REGION Network 28 (STL): spare- VB chan 8
         A     "Epics_to_PLC"."spare-VB-8".cmdSet;
         S     "voie 8 chaufferette BV";
         A     "Epics_to_PLC"."spare-VB-8".cmdRst;
         R     "voie 8 chaufferette BV";
END_REGION

REGION Network 29 (STL): spare- VB chan 9
         A     "Epics_to_PLC"."spare-VB-9".cmdSet;
         S     "voie 9 chaufferette BV";
         A     "Epics_to_PLC"."spare-VB-9".cmdRst;
         R     "voie 9 chaufferette BV";
END_REGION

REGION Network 30 (STL): spare- VB chan 10
         A     "Epics_to_PLC"."spare-VB-10".cmdSet;
         S     "voie 10  chaufferette BV";
         A     "Epics_to_PLC"."spare-VB-10".cmdRst;
         R     "voie 10  chaufferette BV";
END_REGION

REGION Network 31 (STL): spare - VB chan 11
         A     "Epics_to_PLC"."spare-VB-11".cmdSet;
         S     "voie 11 chaufferette BV";
         A     "Epics_to_PLC"."spare-VB-11".cmdRst;
         R     "voie 11 chaufferette BV";
END_REGION

REGION Network 32 (STL): spare - CM chan 5
         A     "Epics_to_PLC"."spare-CM-5".cmdSet;
         S     "voie 5 chaufferette CM";
         A     "Epics_to_PLC"."spare-CM-5".cmdRst;
         R     "voie 5 chaufferette CM";
END_REGION

REGION Network 33 (STL): spare - CM chan 6
         A     "Epics_to_PLC"."spare-CM-6".cmdSet;
         S     "voie 6 chaufferette CM";
         A     "Epics_to_PLC"."spare-CM-6".cmdRst;
         R     "voie 6 chaufferette CM";
END_REGION

REGION Network 34 (STL): spare - CM chan 7
         A     "Epics_to_PLC"."spare-CM-7".cmdSet;
         S     "voie 7 chaufferette CM";
         A     "Epics_to_PLC"."spare-CM-7".cmdRst;
         R     "voie 7 chaufferette CM";
END_REGION

REGION Network 35 (STL): spare - CM chan 8
         A     "Epics_to_PLC"."spare-CM-8".cmdSet;
         S     "voie 8 chaufferette CM";
         A     "Epics_to_PLC"."spare-CM-8".cmdRst;
         R     "voie 8 chaufferette CM";
END_REGION

REGION Network 36 (STL): spare - CM chan 10
         A     "Epics_to_PLC"."spare-CM-10".cmdSet;
         S     "voie 10 chaufferette CM";
         A     "Epics_to_PLC"."spare-CM-10".cmdRst;
         R     "voie 10 chaufferette CM";
END_REGION

REGION Network 37 (STL): spare - CM chan 12
         A     "Epics_to_PLC"."spare-CM-12".cmdSet;
         S     "voie 12 chaufferette CM";
         A     "Epics_to_PLC"."spare-CM-12".cmdRst;
         R     "voie 12 chaufferette CM";
END_REGION

REGION Network 38 (STL): Bit commands
         A     "Epics_to_PLC".cmdAutoMode;
         R     "Graph/manuelle";
         A     "Epics_to_PLC".cmdManMode;
         S     "Graph/manuelle";
         A     "Epics_to_PLC".cmdGrafcetInit;
         =     "MettreEtatInitial";
         A     "Epics_to_PLC".cmdGrafcetErrRst;
         =     "AcquitterErreurGraph";
         A     "Epics_to_PLC".cmdStartConditioning;
         =     "CmdVanneEtatCdt";
         A     "Epics_to_PLC".cmdCondOK;
         =     "CdtInfraOk";
         A     "Epics_to_PLC".cmdCondERR;
         =     "CdtInfraErreur";
         A     "Epics_to_PLC".cmdStartLN2cooling;
         =     "DmdMefAzote";
         A     "Epics_to_PLC".cmdStartLHecooling;
         =     "DmdMefHelium";
         A     "Epics_to_PLC".cmdStart2Kmode;
         =     "DmdMode2K";
         A     "Epics_to_PLC".cmdStop2Kmode;
         =     "DmdArretMode2k";
         A     "Epics_to_PLC".cmdStartSTBYmode;
         =     "DmdModeStandby";
         A     "Epics_to_PLC".cmdStopSTBYmode;
         =     "DmdArretModeStandby";
         A     "Epics_to_PLC".cmdStartHeating;
         =     "StartHeating";
         A     "Epics_to_PLC".cmdStopHeating;
         =     "StopHeating";
         A     "Epics_to_PLC".cmdSelLT01;
         R     "LT_CM".LT02_selCtrl;
         A     "Epics_to_PLC".cmdSelLT02;
         S     "LT_CM".LT02_selCtrl;
END_REGION

REGION Network 39: Real parameters (LHe level PIDs settings)
   RUNG wire#powerrail
      Contact( "Epics_to_PLC".TrigPID_CV01.cmdSet )
      { S7_GenerateENO := "TRUE" } Move(in := "Epics_to_PLC".TrigPID_CV01.cSetV, out1 => "TriggerPIDcv01")
      { S7_GenerateENO := "TRUE" } Move(in := "Epics_to_PLC".TrigPID_CV01.cSetV, out1 => "S8_parameters".TrigPID_CV01)
      R_Coil( "Epics_to_PLC".TrigPID_CV01.cmdSet )
   END_RUNG
   // the same network as SCL:
   // ENO of a box is taken as its EN; it also drops when the box reports an error
   IF "Epics_to_PLC".TrigPID_CV01.cmdSet THEN
       "TriggerPIDcv01" := "Epics_to_PLC".TrigPID_CV01.cSetV;
       "S8_parameters".TrigPID_CV01 := "Epics_to_PLC".TrigPID_CV01.cSetV;
       "Epics_to_PLC".TrigPID_CV01.cmdSet := FALSE;
   END_IF;
END_REGION

REGION Network 40: Real parameters (LHe level PIDs settings)
   RUNG wire#powerrail
      Contact( "Epics_to_PLC".TrigPID_CV02.cmdSet )
      { S7_GenerateENO := "TRUE" } Move(in := "Epics_to_PLC".TrigPID_CV02.cSetV, out1 => "TriggerPIDcv02")
      { S7_GenerateENO := "TRUE" } Move(in := "Epics_to_PLC".TrigPID_CV02.cSetV, out1 => "S6_parameters".TrigPID_CV02)
      R_Coil( "Epics_to_PLC".TrigPID_CV02.cmdSet )
   END_RUNG
   // the same network as SCL:
   // ENO of a box is taken as its EN; it also drops when the box reports an error
   IF "Epics_to_PLC".TrigPID_CV02.cmdSet THEN
       "TriggerPIDcv02" := "Epics_to_PLC".TrigPID_CV02.cSetV;
       "S6_parameters".TrigPID_CV02 := "Epics_to_PLC".TrigPID_CV02.cSetV;
       "Epics_to_PLC".TrigPID_CV02.cmdSet := FALSE;
   END_IF;
END_REGION

REGION Network 41: Real parameters (LHe level PIDs settings)
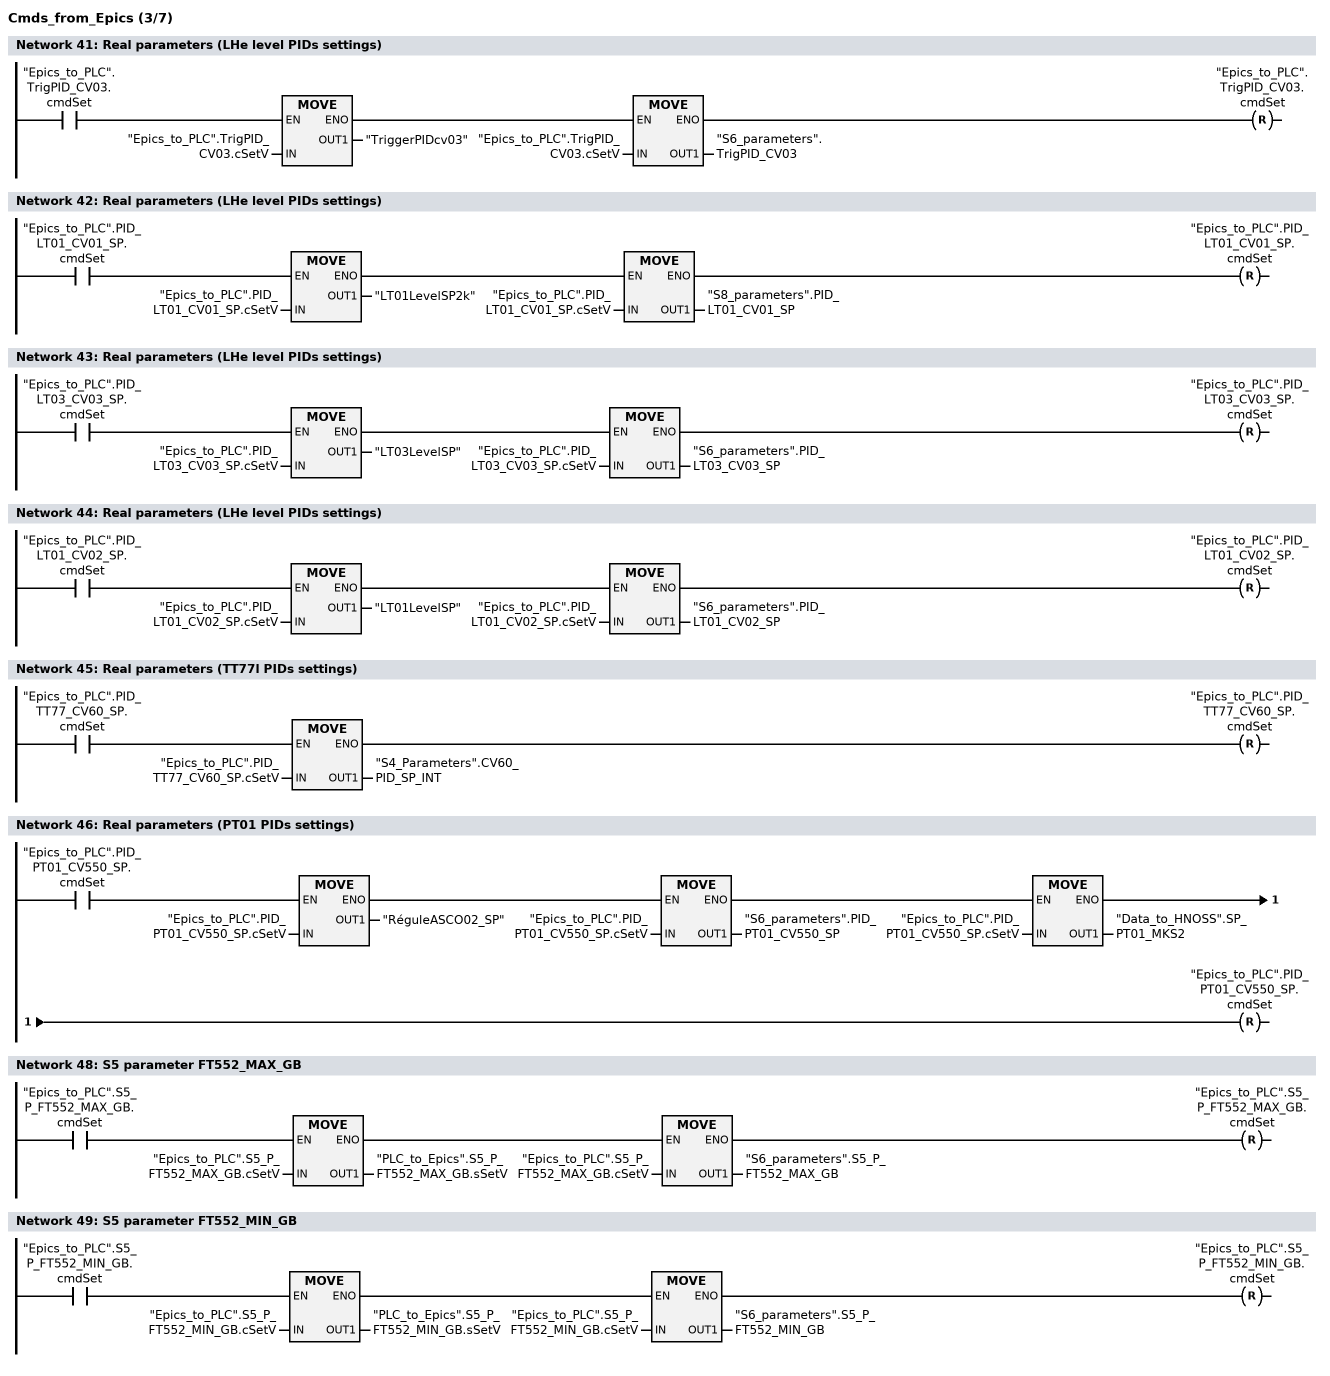
   RUNG wire#powerrail
      Contact( "Epics_to_PLC".TrigPID_CV03.cmdSet )
      { S7_GenerateENO := "TRUE" } Move(in := "Epics_to_PLC".TrigPID_CV03.cSetV, out1 => "TriggerPIDcv03")
      { S7_GenerateENO := "TRUE" } Move(in := "Epics_to_PLC".TrigPID_CV03.cSetV, out1 => "S6_parameters".TrigPID_CV03)
      R_Coil( "Epics_to_PLC".TrigPID_CV03.cmdSet )
   END_RUNG
   // the same network as SCL:
   // ENO of a box is taken as its EN; it also drops when the box reports an error
   IF "Epics_to_PLC".TrigPID_CV03.cmdSet THEN
       "TriggerPIDcv03" := "Epics_to_PLC".TrigPID_CV03.cSetV;
       "S6_parameters".TrigPID_CV03 := "Epics_to_PLC".TrigPID_CV03.cSetV;
       "Epics_to_PLC".TrigPID_CV03.cmdSet := FALSE;
   END_IF;
END_REGION

REGION Network 42: Real parameters (LHe level PIDs settings)
   RUNG wire#powerrail
      Contact( "Epics_to_PLC".PID_LT01_CV01_SP.cmdSet )
      { S7_GenerateENO := "TRUE" } Move(in := "Epics_to_PLC".PID_LT01_CV01_SP.cSetV, out1 => "LT01LevelSP2k")
      { S7_GenerateENO := "TRUE" } Move(in := "Epics_to_PLC".PID_LT01_CV01_SP.cSetV, out1 => "S8_parameters".PID_LT01_CV01_SP)
      R_Coil( "Epics_to_PLC".PID_LT01_CV01_SP.cmdSet )
   END_RUNG
   // the same network as SCL:
   // ENO of a box is taken as its EN; it also drops when the box reports an error
   IF "Epics_to_PLC".PID_LT01_CV01_SP.cmdSet THEN
       "LT01LevelSP2k" := "Epics_to_PLC".PID_LT01_CV01_SP.cSetV;
       "S8_parameters".PID_LT01_CV01_SP := "Epics_to_PLC".PID_LT01_CV01_SP.cSetV;
       "Epics_to_PLC".PID_LT01_CV01_SP.cmdSet := FALSE;
   END_IF;
END_REGION

REGION Network 43: Real parameters (LHe level PIDs settings)
   RUNG wire#powerrail
      Contact( "Epics_to_PLC".PID_LT03_CV03_SP.cmdSet )
      { S7_GenerateENO := "TRUE" } Move(in := "Epics_to_PLC".PID_LT03_CV03_SP.cSetV, out1 => "LT03LevelSP")
      { S7_GenerateENO := "TRUE" } Move(in := "Epics_to_PLC".PID_LT03_CV03_SP.cSetV, out1 => "S6_parameters".PID_LT03_CV03_SP)
      R_Coil( "Epics_to_PLC".PID_LT03_CV03_SP.cmdSet )
   END_RUNG
   // the same network as SCL:
   // ENO of a box is taken as its EN; it also drops when the box reports an error
   IF "Epics_to_PLC".PID_LT03_CV03_SP.cmdSet THEN
       "LT03LevelSP" := "Epics_to_PLC".PID_LT03_CV03_SP.cSetV;
       "S6_parameters".PID_LT03_CV03_SP := "Epics_to_PLC".PID_LT03_CV03_SP.cSetV;
       "Epics_to_PLC".PID_LT03_CV03_SP.cmdSet := FALSE;
   END_IF;
END_REGION

REGION Network 44: Real parameters (LHe level PIDs settings)
   RUNG wire#powerrail
      Contact( "Epics_to_PLC".PID_LT01_CV02_SP.cmdSet )
      { S7_GenerateENO := "TRUE" } Move(in := "Epics_to_PLC".PID_LT01_CV02_SP.cSetV, out1 => "LT01LevelSP")
      { S7_GenerateENO := "TRUE" } Move(in := "Epics_to_PLC".PID_LT01_CV02_SP.cSetV, out1 => "S6_parameters".PID_LT01_CV02_SP)
      R_Coil( "Epics_to_PLC".PID_LT01_CV02_SP.cmdSet )
   END_RUNG
   // the same network as SCL:
   // ENO of a box is taken as its EN; it also drops when the box reports an error
   IF "Epics_to_PLC".PID_LT01_CV02_SP.cmdSet THEN
       "LT01LevelSP" := "Epics_to_PLC".PID_LT01_CV02_SP.cSetV;
       "S6_parameters".PID_LT01_CV02_SP := "Epics_to_PLC".PID_LT01_CV02_SP.cSetV;
       "Epics_to_PLC".PID_LT01_CV02_SP.cmdSet := FALSE;
   END_IF;
END_REGION

REGION Network 45: Real parameters (TT77l PIDs settings)
   RUNG wire#powerrail
      Contact( "Epics_to_PLC".PID_TT77_CV60_SP.cmdSet )
      { S7_GenerateENO := "TRUE" } Move(in := "Epics_to_PLC".PID_TT77_CV60_SP.cSetV, out1 => "S4_Parameters".CV60_PID_SP_INT)
      R_Coil( "Epics_to_PLC".PID_TT77_CV60_SP.cmdSet )
   END_RUNG
   // the same network as SCL:
   // ENO of a box is taken as its EN; it also drops when the box reports an error
   IF "Epics_to_PLC".PID_TT77_CV60_SP.cmdSet THEN
       "S4_Parameters".CV60_PID_SP_INT := "Epics_to_PLC".PID_TT77_CV60_SP.cSetV;
       "Epics_to_PLC".PID_TT77_CV60_SP.cmdSet := FALSE;
   END_IF;
END_REGION

REGION Network 46: Real parameters (PT01 PIDs settings)
   RUNG wire#powerrail
      Contact( "Epics_to_PLC".PID_PT01_CV550_SP.cmdSet )
      { S7_GenerateENO := "TRUE" } Move(in := "Epics_to_PLC".PID_PT01_CV550_SP.cSetV, out1 => "RéguleASCO02_SP")
      { S7_GenerateENO := "TRUE" } Move(in := "Epics_to_PLC".PID_PT01_CV550_SP.cSetV, out1 => "S6_parameters".PID_PT01_CV550_SP)
      { S7_GenerateENO := "TRUE" } Move(in := "Epics_to_PLC".PID_PT01_CV550_SP.cSetV, out1 => "Data_to_HNOSS".SP_PT01_MKS2)
      R_Coil( "Epics_to_PLC".PID_PT01_CV550_SP.cmdSet )
   END_RUNG
   // the same network as SCL:
   // ENO of a box is taken as its EN; it also drops when the box reports an error
   IF "Epics_to_PLC".PID_PT01_CV550_SP.cmdSet THEN
       "RéguleASCO02_SP" := "Epics_to_PLC".PID_PT01_CV550_SP.cSetV;
       "S6_parameters".PID_PT01_CV550_SP := "Epics_to_PLC".PID_PT01_CV550_SP.cSetV;
       "Data_to_HNOSS".SP_PT01_MKS2 := "Epics_to_PLC".PID_PT01_CV550_SP.cSetV;
       "Epics_to_PLC".PID_PT01_CV550_SP.cmdSet := FALSE;
   END_IF;
END_REGION

REGION Network 47 (STL): Temperatures fromKeithley
         L     "Epics_to_PLC".TTxx;
         T     "ReceivePT100"."TTxx_(K)";
         L     "Epics_to_PLC".TTyy;
         T     "ReceivePT100"."TTyy_(K)";
END_REGION

REGION Network 48: S5 parameter FT552_MAX_GB
   RUNG wire#powerrail
      Contact( "Epics_to_PLC".S5_P_FT552_MAX_GB.cmdSet )
      { S7_GenerateENO := "TRUE" } Move(in := "Epics_to_PLC".S5_P_FT552_MAX_GB.cSetV, out1 => "PLC_to_Epics".S5_P_FT552_MAX_GB.sSetV)
      { S7_GenerateENO := "TRUE" } Move(in := "Epics_to_PLC".S5_P_FT552_MAX_GB.cSetV, out1 => "S6_parameters".S5_P_FT552_MAX_GB)
      R_Coil( "Epics_to_PLC".S5_P_FT552_MAX_GB.cmdSet )
   END_RUNG
   // the same network as SCL:
   // ENO of a box is taken as its EN; it also drops when the box reports an error
   IF "Epics_to_PLC".S5_P_FT552_MAX_GB.cmdSet THEN
       "PLC_to_Epics".S5_P_FT552_MAX_GB.sSetV := "Epics_to_PLC".S5_P_FT552_MAX_GB.cSetV;
       "S6_parameters".S5_P_FT552_MAX_GB := "Epics_to_PLC".S5_P_FT552_MAX_GB.cSetV;
       "Epics_to_PLC".S5_P_FT552_MAX_GB.cmdSet := FALSE;
   END_IF;
END_REGION

REGION Network 49: S5 parameter FT552_MIN_GB
   RUNG wire#powerrail
      Contact( "Epics_to_PLC".S5_P_FT552_MIN_GB.cmdSet )
      { S7_GenerateENO := "TRUE" } Move(in := "Epics_to_PLC".S5_P_FT552_MIN_GB.cSetV, out1 => "PLC_to_Epics".S5_P_FT552_MIN_GB.sSetV)
      { S7_GenerateENO := "TRUE" } Move(in := "Epics_to_PLC".S5_P_FT552_MIN_GB.cSetV, out1 => "S6_parameters".S5_P_FT552_MIN_GB)
      R_Coil( "Epics_to_PLC".S5_P_FT552_MIN_GB.cmdSet )
   END_RUNG
   // the same network as SCL:
   // ENO of a box is taken as its EN; it also drops when the box reports an error
   IF "Epics_to_PLC".S5_P_FT552_MIN_GB.cmdSet THEN
       "PLC_to_Epics".S5_P_FT552_MIN_GB.sSetV := "Epics_to_PLC".S5_P_FT552_MIN_GB.cSetV;
       "S6_parameters".S5_P_FT552_MIN_GB := "Epics_to_PLC".S5_P_FT552_MIN_GB.cSetV;
       "Epics_to_PLC".S5_P_FT552_MIN_GB.cmdSet := FALSE;
   END_IF;
END_REGION

REGION Network 50: S5 parameter FT552_MAX_C
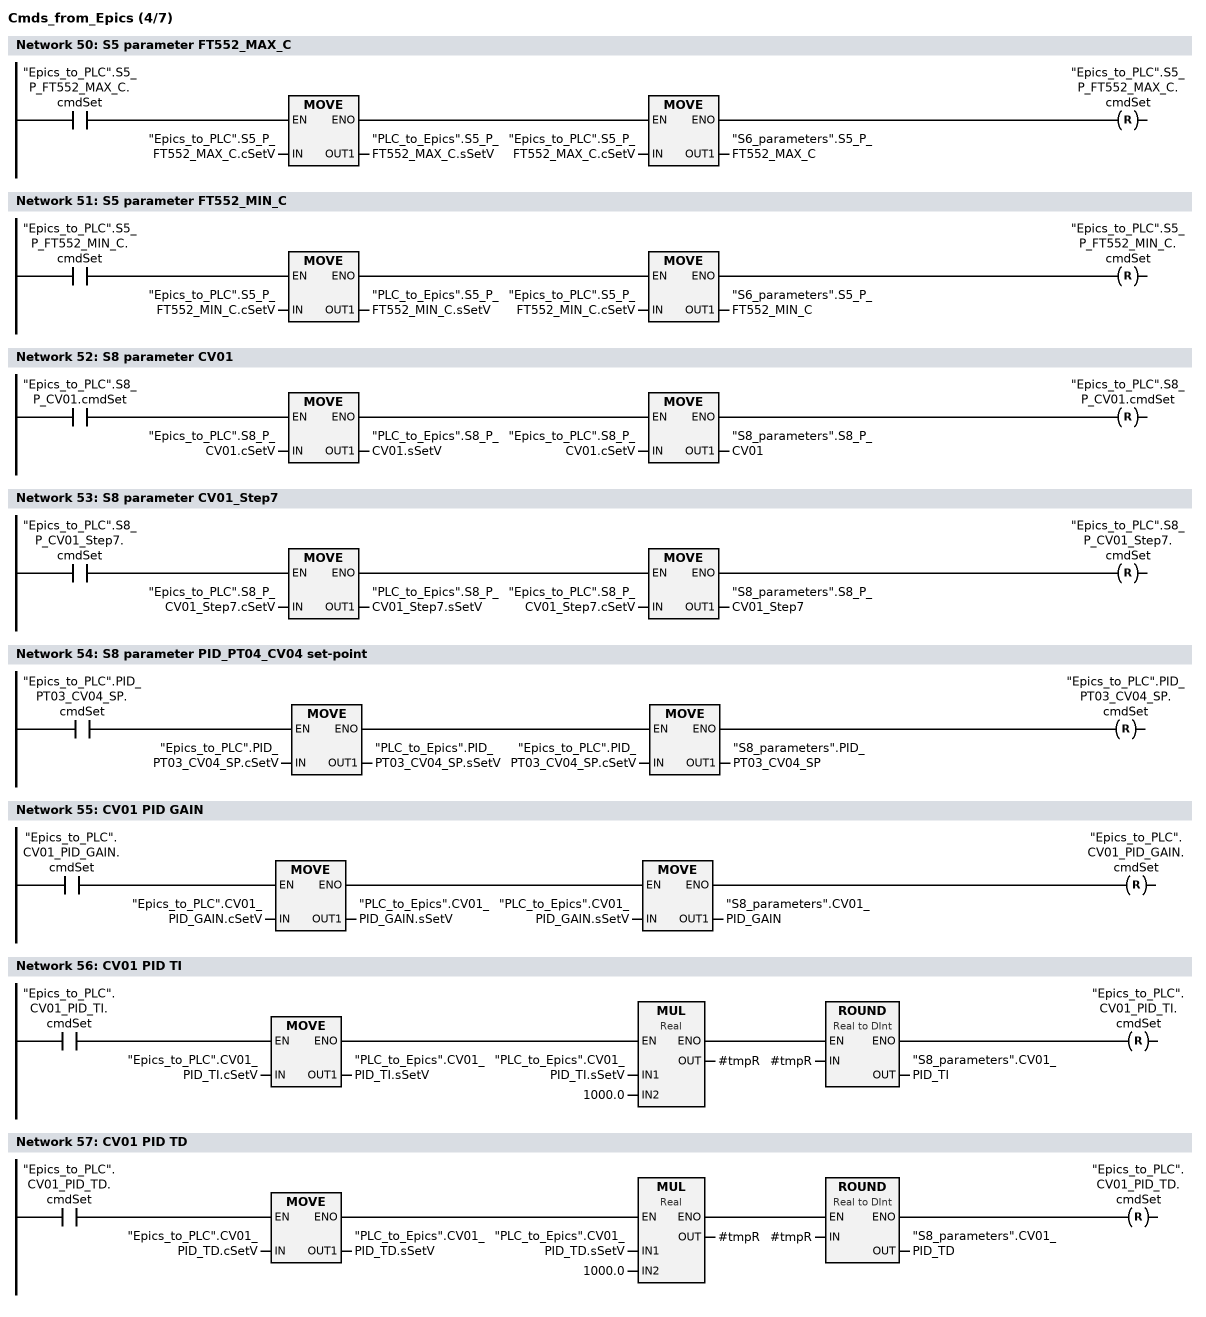
   RUNG wire#powerrail
      Contact( "Epics_to_PLC".S5_P_FT552_MAX_C.cmdSet )
      { S7_GenerateENO := "TRUE" } Move(in := "Epics_to_PLC".S5_P_FT552_MAX_C.cSetV, out1 => "PLC_to_Epics".S5_P_FT552_MAX_C.sSetV)
      { S7_GenerateENO := "TRUE" } Move(in := "Epics_to_PLC".S5_P_FT552_MAX_C.cSetV, out1 => "S6_parameters".S5_P_FT552_MAX_C)
      R_Coil( "Epics_to_PLC".S5_P_FT552_MAX_C.cmdSet )
   END_RUNG
   // the same network as SCL:
   // ENO of a box is taken as its EN; it also drops when the box reports an error
   IF "Epics_to_PLC".S5_P_FT552_MAX_C.cmdSet THEN
       "PLC_to_Epics".S5_P_FT552_MAX_C.sSetV := "Epics_to_PLC".S5_P_FT552_MAX_C.cSetV;
       "S6_parameters".S5_P_FT552_MAX_C := "Epics_to_PLC".S5_P_FT552_MAX_C.cSetV;
       "Epics_to_PLC".S5_P_FT552_MAX_C.cmdSet := FALSE;
   END_IF;
END_REGION

REGION Network 51: S5 parameter FT552_MIN_C
   RUNG wire#powerrail
      Contact( "Epics_to_PLC".S5_P_FT552_MIN_C.cmdSet )
      { S7_GenerateENO := "TRUE" } Move(in := "Epics_to_PLC".S5_P_FT552_MIN_C.cSetV, out1 => "PLC_to_Epics".S5_P_FT552_MIN_C.sSetV)
      { S7_GenerateENO := "TRUE" } Move(in := "Epics_to_PLC".S5_P_FT552_MIN_C.cSetV, out1 => "S6_parameters".S5_P_FT552_MIN_C)
      R_Coil( "Epics_to_PLC".S5_P_FT552_MIN_C.cmdSet )
   END_RUNG
   // the same network as SCL:
   // ENO of a box is taken as its EN; it also drops when the box reports an error
   IF "Epics_to_PLC".S5_P_FT552_MIN_C.cmdSet THEN
       "PLC_to_Epics".S5_P_FT552_MIN_C.sSetV := "Epics_to_PLC".S5_P_FT552_MIN_C.cSetV;
       "S6_parameters".S5_P_FT552_MIN_C := "Epics_to_PLC".S5_P_FT552_MIN_C.cSetV;
       "Epics_to_PLC".S5_P_FT552_MIN_C.cmdSet := FALSE;
   END_IF;
END_REGION

REGION Network 52: S8 parameter CV01
   RUNG wire#powerrail
      Contact( "Epics_to_PLC".S8_P_CV01.cmdSet )
      { S7_GenerateENO := "TRUE" } Move(in := "Epics_to_PLC".S8_P_CV01.cSetV, out1 => "PLC_to_Epics".S8_P_CV01.sSetV)
      { S7_GenerateENO := "TRUE" } Move(in := "Epics_to_PLC".S8_P_CV01.cSetV, out1 => "S8_parameters".S8_P_CV01)
      R_Coil( "Epics_to_PLC".S8_P_CV01.cmdSet )
   END_RUNG
   // the same network as SCL:
   // ENO of a box is taken as its EN; it also drops when the box reports an error
   IF "Epics_to_PLC".S8_P_CV01.cmdSet THEN
       "PLC_to_Epics".S8_P_CV01.sSetV := "Epics_to_PLC".S8_P_CV01.cSetV;
       "S8_parameters".S8_P_CV01 := "Epics_to_PLC".S8_P_CV01.cSetV;
       "Epics_to_PLC".S8_P_CV01.cmdSet := FALSE;
   END_IF;
END_REGION

REGION Network 53: S8 parameter CV01_Step7
   RUNG wire#powerrail
      Contact( "Epics_to_PLC".S8_P_CV01_Step7.cmdSet )
      { S7_GenerateENO := "TRUE" } Move(in := "Epics_to_PLC".S8_P_CV01_Step7.cSetV, out1 => "PLC_to_Epics".S8_P_CV01_Step7.sSetV)
      { S7_GenerateENO := "TRUE" } Move(in := "Epics_to_PLC".S8_P_CV01_Step7.cSetV, out1 => "S8_parameters".S8_P_CV01_Step7)
      R_Coil( "Epics_to_PLC".S8_P_CV01_Step7.cmdSet )
   END_RUNG
   // the same network as SCL:
   // ENO of a box is taken as its EN; it also drops when the box reports an error
   IF "Epics_to_PLC".S8_P_CV01_Step7.cmdSet THEN
       "PLC_to_Epics".S8_P_CV01_Step7.sSetV := "Epics_to_PLC".S8_P_CV01_Step7.cSetV;
       "S8_parameters".S8_P_CV01_Step7 := "Epics_to_PLC".S8_P_CV01_Step7.cSetV;
       "Epics_to_PLC".S8_P_CV01_Step7.cmdSet := FALSE;
   END_IF;
END_REGION

REGION Network 54: S8 parameter PID_PT04_CV04 set-point
   RUNG wire#powerrail
      Contact( "Epics_to_PLC".PID_PT03_CV04_SP.cmdSet )
      { S7_GenerateENO := "TRUE" } Move(in := "Epics_to_PLC".PID_PT03_CV04_SP.cSetV, out1 => "PLC_to_Epics".PID_PT03_CV04_SP.sSetV)
      { S7_GenerateENO := "TRUE" } Move(in := "Epics_to_PLC".PID_PT03_CV04_SP.cSetV, out1 => "S8_parameters".PID_PT03_CV04_SP)
      R_Coil( "Epics_to_PLC".PID_PT03_CV04_SP.cmdSet )
   END_RUNG
   // the same network as SCL:
   // ENO of a box is taken as its EN; it also drops when the box reports an error
   IF "Epics_to_PLC".PID_PT03_CV04_SP.cmdSet THEN
       "PLC_to_Epics".PID_PT03_CV04_SP.sSetV := "Epics_to_PLC".PID_PT03_CV04_SP.cSetV;
       "S8_parameters".PID_PT03_CV04_SP := "Epics_to_PLC".PID_PT03_CV04_SP.cSetV;
       "Epics_to_PLC".PID_PT03_CV04_SP.cmdSet := FALSE;
   END_IF;
END_REGION

REGION Network 55: CV01 PID GAIN
   RUNG wire#powerrail
      Contact( "Epics_to_PLC".CV01_PID_GAIN.cmdSet )
      { S7_GenerateENO := "TRUE" } Move(in := "Epics_to_PLC".CV01_PID_GAIN.cSetV, out1 => "PLC_to_Epics".CV01_PID_GAIN.sSetV)
      { S7_GenerateENO := "TRUE" } Move(in := "PLC_to_Epics".CV01_PID_GAIN.sSetV, out1 => "S8_parameters".CV01_PID_GAIN)
      R_Coil( "Epics_to_PLC".CV01_PID_GAIN.cmdSet )
   END_RUNG
   // the same network as SCL:
   // ENO of a box is taken as its EN; it also drops when the box reports an error
   IF "Epics_to_PLC".CV01_PID_GAIN.cmdSet THEN
       "PLC_to_Epics".CV01_PID_GAIN.sSetV := "Epics_to_PLC".CV01_PID_GAIN.cSetV;
       "S8_parameters".CV01_PID_GAIN := "PLC_to_Epics".CV01_PID_GAIN.sSetV;
       "Epics_to_PLC".CV01_PID_GAIN.cmdSet := FALSE;
   END_IF;
END_REGION

REGION Network 56: CV01 PID TI
   RUNG wire#powerrail
      Contact( "Epics_to_PLC".CV01_PID_TI.cmdSet )
      { S7_GenerateENO := "TRUE" } Move(in := "Epics_to_PLC".CV01_PID_TI.cSetV, out1 => "PLC_to_Epics".CV01_PID_TI.sSetV)
      { S7_Templates := "SrcType := Real"; S7_GenerateENO := "TRUE" } Mul(in1 := "PLC_to_Epics".CV01_PID_TI.sSetV, in2 := 1000.0, out => #tmpR)
      { S7_Templates := "[SrcType := Real, DestType := DInt]"; S7_GenerateENO := "TRUE" } Round(in := #tmpR, out => "S8_parameters".CV01_PID_TI)
      R_Coil( "Epics_to_PLC".CV01_PID_TI.cmdSet )
   END_RUNG
   // the same network as SCL:
   // ENO of a box is taken as its EN; it also drops when the box reports an error
   IF "Epics_to_PLC".CV01_PID_TI.cmdSet THEN
       "PLC_to_Epics".CV01_PID_TI.sSetV := "Epics_to_PLC".CV01_PID_TI.cSetV;
       #tmpR := "PLC_to_Epics".CV01_PID_TI.sSetV * 1000.0;
       "S8_parameters".CV01_PID_TI := ROUND(#tmpR);
       "Epics_to_PLC".CV01_PID_TI.cmdSet := FALSE;
   END_IF;
END_REGION

REGION Network 57: CV01 PID TD
   RUNG wire#powerrail
      Contact( "Epics_to_PLC".CV01_PID_TD.cmdSet )
      { S7_GenerateENO := "TRUE" } Move(in := "Epics_to_PLC".CV01_PID_TD.cSetV, out1 => "PLC_to_Epics".CV01_PID_TD.sSetV)
      { S7_Templates := "SrcType := Real"; S7_GenerateENO := "TRUE" } Mul(in1 := "PLC_to_Epics".CV01_PID_TD.sSetV, in2 := 1000.0, out => #tmpR)
      { S7_Templates := "[SrcType := Real, DestType := DInt]"; S7_GenerateENO := "TRUE" } Round(in := #tmpR, out => "S8_parameters".CV01_PID_TD)
      R_Coil( "Epics_to_PLC".CV01_PID_TD.cmdSet )
   END_RUNG
   // the same network as SCL:
   // ENO of a box is taken as its EN; it also drops when the box reports an error
   IF "Epics_to_PLC".CV01_PID_TD.cmdSet THEN
       "PLC_to_Epics".CV01_PID_TD.sSetV := "Epics_to_PLC".CV01_PID_TD.cSetV;
       #tmpR := "PLC_to_Epics".CV01_PID_TD.sSetV * 1000.0;
       "S8_parameters".CV01_PID_TD := ROUND(#tmpR);
       "Epics_to_PLC".CV01_PID_TD.cmdSet := FALSE;
   END_IF;
END_REGION

REGION Network 58: CV01 PID TM_LAG
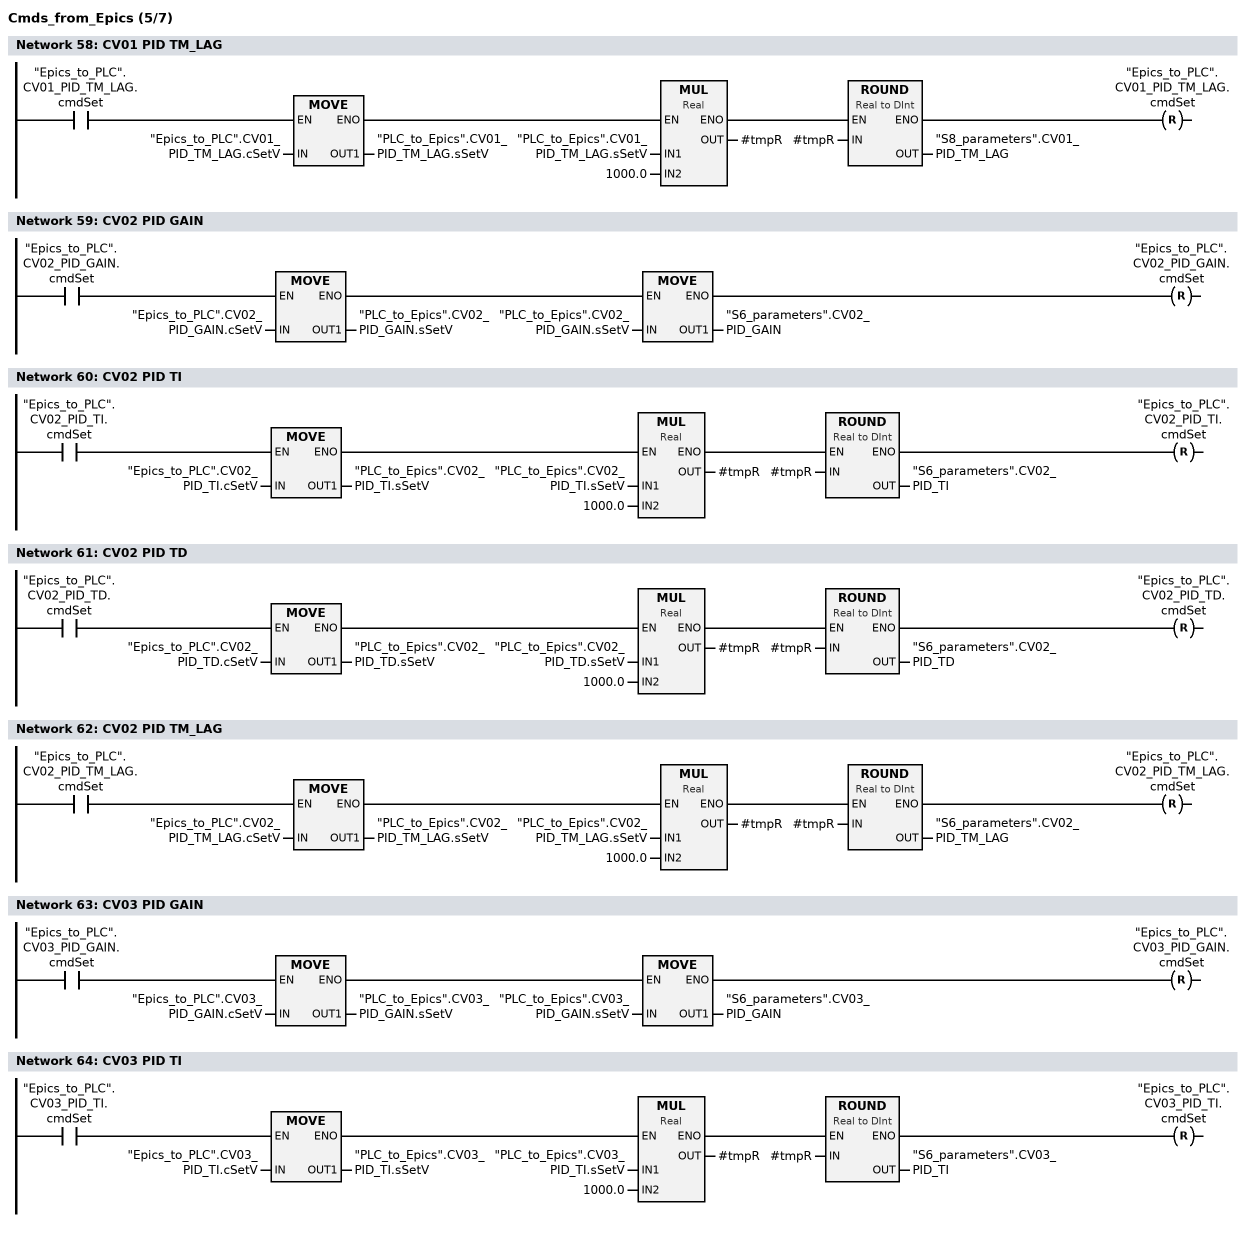
   RUNG wire#powerrail
      Contact( "Epics_to_PLC".CV01_PID_TM_LAG.cmdSet )
      { S7_GenerateENO := "TRUE" } Move(in := "Epics_to_PLC".CV01_PID_TM_LAG.cSetV, out1 => "PLC_to_Epics".CV01_PID_TM_LAG.sSetV)
      { S7_Templates := "SrcType := Real"; S7_GenerateENO := "TRUE" } Mul(in1 := "PLC_to_Epics".CV01_PID_TM_LAG.sSetV, in2 := 1000.0, out => #tmpR)
      { S7_Templates := "[SrcType := Real, DestType := DInt]"; S7_GenerateENO := "TRUE" } Round(in := #tmpR, out => "S8_parameters".CV01_PID_TM_LAG)
      R_Coil( "Epics_to_PLC".CV01_PID_TM_LAG.cmdSet )
   END_RUNG
   // the same network as SCL:
   // ENO of a box is taken as its EN; it also drops when the box reports an error
   IF "Epics_to_PLC".CV01_PID_TM_LAG.cmdSet THEN
       "PLC_to_Epics".CV01_PID_TM_LAG.sSetV := "Epics_to_PLC".CV01_PID_TM_LAG.cSetV;
       #tmpR := "PLC_to_Epics".CV01_PID_TM_LAG.sSetV * 1000.0;
       "S8_parameters".CV01_PID_TM_LAG := ROUND(#tmpR);
       "Epics_to_PLC".CV01_PID_TM_LAG.cmdSet := FALSE;
   END_IF;
END_REGION

REGION Network 59: CV02 PID GAIN
   RUNG wire#powerrail
      Contact( "Epics_to_PLC".CV02_PID_GAIN.cmdSet )
      { S7_GenerateENO := "TRUE" } Move(in := "Epics_to_PLC".CV02_PID_GAIN.cSetV, out1 => "PLC_to_Epics".CV02_PID_GAIN.sSetV)
      { S7_GenerateENO := "TRUE" } Move(in := "PLC_to_Epics".CV02_PID_GAIN.sSetV, out1 => "S6_parameters".CV02_PID_GAIN)
      R_Coil( "Epics_to_PLC".CV02_PID_GAIN.cmdSet )
   END_RUNG
   // the same network as SCL:
   // ENO of a box is taken as its EN; it also drops when the box reports an error
   IF "Epics_to_PLC".CV02_PID_GAIN.cmdSet THEN
       "PLC_to_Epics".CV02_PID_GAIN.sSetV := "Epics_to_PLC".CV02_PID_GAIN.cSetV;
       "S6_parameters".CV02_PID_GAIN := "PLC_to_Epics".CV02_PID_GAIN.sSetV;
       "Epics_to_PLC".CV02_PID_GAIN.cmdSet := FALSE;
   END_IF;
END_REGION

REGION Network 60: CV02 PID TI
   RUNG wire#powerrail
      Contact( "Epics_to_PLC".CV02_PID_TI.cmdSet )
      { S7_GenerateENO := "TRUE" } Move(in := "Epics_to_PLC".CV02_PID_TI.cSetV, out1 => "PLC_to_Epics".CV02_PID_TI.sSetV)
      { S7_Templates := "SrcType := Real"; S7_GenerateENO := "TRUE" } Mul(in1 := "PLC_to_Epics".CV02_PID_TI.sSetV, in2 := 1000.0, out => #tmpR)
      { S7_Templates := "[SrcType := Real, DestType := DInt]"; S7_GenerateENO := "TRUE" } Round(in := #tmpR, out => "S6_parameters".CV02_PID_TI)
      R_Coil( "Epics_to_PLC".CV02_PID_TI.cmdSet )
   END_RUNG
   // the same network as SCL:
   // ENO of a box is taken as its EN; it also drops when the box reports an error
   IF "Epics_to_PLC".CV02_PID_TI.cmdSet THEN
       "PLC_to_Epics".CV02_PID_TI.sSetV := "Epics_to_PLC".CV02_PID_TI.cSetV;
       #tmpR := "PLC_to_Epics".CV02_PID_TI.sSetV * 1000.0;
       "S6_parameters".CV02_PID_TI := ROUND(#tmpR);
       "Epics_to_PLC".CV02_PID_TI.cmdSet := FALSE;
   END_IF;
END_REGION

REGION Network 61: CV02 PID TD
   RUNG wire#powerrail
      Contact( "Epics_to_PLC".CV02_PID_TD.cmdSet )
      { S7_GenerateENO := "TRUE" } Move(in := "Epics_to_PLC".CV02_PID_TD.cSetV, out1 => "PLC_to_Epics".CV02_PID_TD.sSetV)
      { S7_Templates := "SrcType := Real"; S7_GenerateENO := "TRUE" } Mul(in1 := "PLC_to_Epics".CV02_PID_TD.sSetV, in2 := 1000.0, out => #tmpR)
      { S7_Templates := "[SrcType := Real, DestType := DInt]"; S7_GenerateENO := "TRUE" } Round(in := #tmpR, out => "S6_parameters".CV02_PID_TD)
      R_Coil( "Epics_to_PLC".CV02_PID_TD.cmdSet )
   END_RUNG
   // the same network as SCL:
   // ENO of a box is taken as its EN; it also drops when the box reports an error
   IF "Epics_to_PLC".CV02_PID_TD.cmdSet THEN
       "PLC_to_Epics".CV02_PID_TD.sSetV := "Epics_to_PLC".CV02_PID_TD.cSetV;
       #tmpR := "PLC_to_Epics".CV02_PID_TD.sSetV * 1000.0;
       "S6_parameters".CV02_PID_TD := ROUND(#tmpR);
       "Epics_to_PLC".CV02_PID_TD.cmdSet := FALSE;
   END_IF;
END_REGION

REGION Network 62: CV02 PID TM_LAG
   RUNG wire#powerrail
      Contact( "Epics_to_PLC".CV02_PID_TM_LAG.cmdSet )
      { S7_GenerateENO := "TRUE" } Move(in := "Epics_to_PLC".CV02_PID_TM_LAG.cSetV, out1 => "PLC_to_Epics".CV02_PID_TM_LAG.sSetV)
      { S7_Templates := "SrcType := Real"; S7_GenerateENO := "TRUE" } Mul(in1 := "PLC_to_Epics".CV02_PID_TM_LAG.sSetV, in2 := 1000.0, out => #tmpR)
      { S7_Templates := "[SrcType := Real, DestType := DInt]"; S7_GenerateENO := "TRUE" } Round(in := #tmpR, out => "S6_parameters".CV02_PID_TM_LAG)
      R_Coil( "Epics_to_PLC".CV02_PID_TM_LAG.cmdSet )
   END_RUNG
   // the same network as SCL:
   // ENO of a box is taken as its EN; it also drops when the box reports an error
   IF "Epics_to_PLC".CV02_PID_TM_LAG.cmdSet THEN
       "PLC_to_Epics".CV02_PID_TM_LAG.sSetV := "Epics_to_PLC".CV02_PID_TM_LAG.cSetV;
       #tmpR := "PLC_to_Epics".CV02_PID_TM_LAG.sSetV * 1000.0;
       "S6_parameters".CV02_PID_TM_LAG := ROUND(#tmpR);
       "Epics_to_PLC".CV02_PID_TM_LAG.cmdSet := FALSE;
   END_IF;
END_REGION

REGION Network 63: CV03 PID GAIN
   RUNG wire#powerrail
      Contact( "Epics_to_PLC".CV03_PID_GAIN.cmdSet )
      { S7_GenerateENO := "TRUE" } Move(in := "Epics_to_PLC".CV03_PID_GAIN.cSetV, out1 => "PLC_to_Epics".CV03_PID_GAIN.sSetV)
      { S7_GenerateENO := "TRUE" } Move(in := "PLC_to_Epics".CV03_PID_GAIN.sSetV, out1 => "S6_parameters".CV03_PID_GAIN)
      R_Coil( "Epics_to_PLC".CV03_PID_GAIN.cmdSet )
   END_RUNG
   // the same network as SCL:
   // ENO of a box is taken as its EN; it also drops when the box reports an error
   IF "Epics_to_PLC".CV03_PID_GAIN.cmdSet THEN
       "PLC_to_Epics".CV03_PID_GAIN.sSetV := "Epics_to_PLC".CV03_PID_GAIN.cSetV;
       "S6_parameters".CV03_PID_GAIN := "PLC_to_Epics".CV03_PID_GAIN.sSetV;
       "Epics_to_PLC".CV03_PID_GAIN.cmdSet := FALSE;
   END_IF;
END_REGION

REGION Network 64: CV03 PID TI
   RUNG wire#powerrail
      Contact( "Epics_to_PLC".CV03_PID_TI.cmdSet )
      { S7_GenerateENO := "TRUE" } Move(in := "Epics_to_PLC".CV03_PID_TI.cSetV, out1 => "PLC_to_Epics".CV03_PID_TI.sSetV)
      { S7_Templates := "SrcType := Real"; S7_GenerateENO := "TRUE" } Mul(in1 := "PLC_to_Epics".CV03_PID_TI.sSetV, in2 := 1000.0, out => #tmpR)
      { S7_Templates := "[SrcType := Real, DestType := DInt]"; S7_GenerateENO := "TRUE" } Round(in := #tmpR, out => "S6_parameters".CV03_PID_TI)
      R_Coil( "Epics_to_PLC".CV03_PID_TI.cmdSet )
   END_RUNG
   // the same network as SCL:
   // ENO of a box is taken as its EN; it also drops when the box reports an error
   IF "Epics_to_PLC".CV03_PID_TI.cmdSet THEN
       "PLC_to_Epics".CV03_PID_TI.sSetV := "Epics_to_PLC".CV03_PID_TI.cSetV;
       #tmpR := "PLC_to_Epics".CV03_PID_TI.sSetV * 1000.0;
       "S6_parameters".CV03_PID_TI := ROUND(#tmpR);
       "Epics_to_PLC".CV03_PID_TI.cmdSet := FALSE;
   END_IF;
END_REGION

REGION Network 65: CV03 PID TD
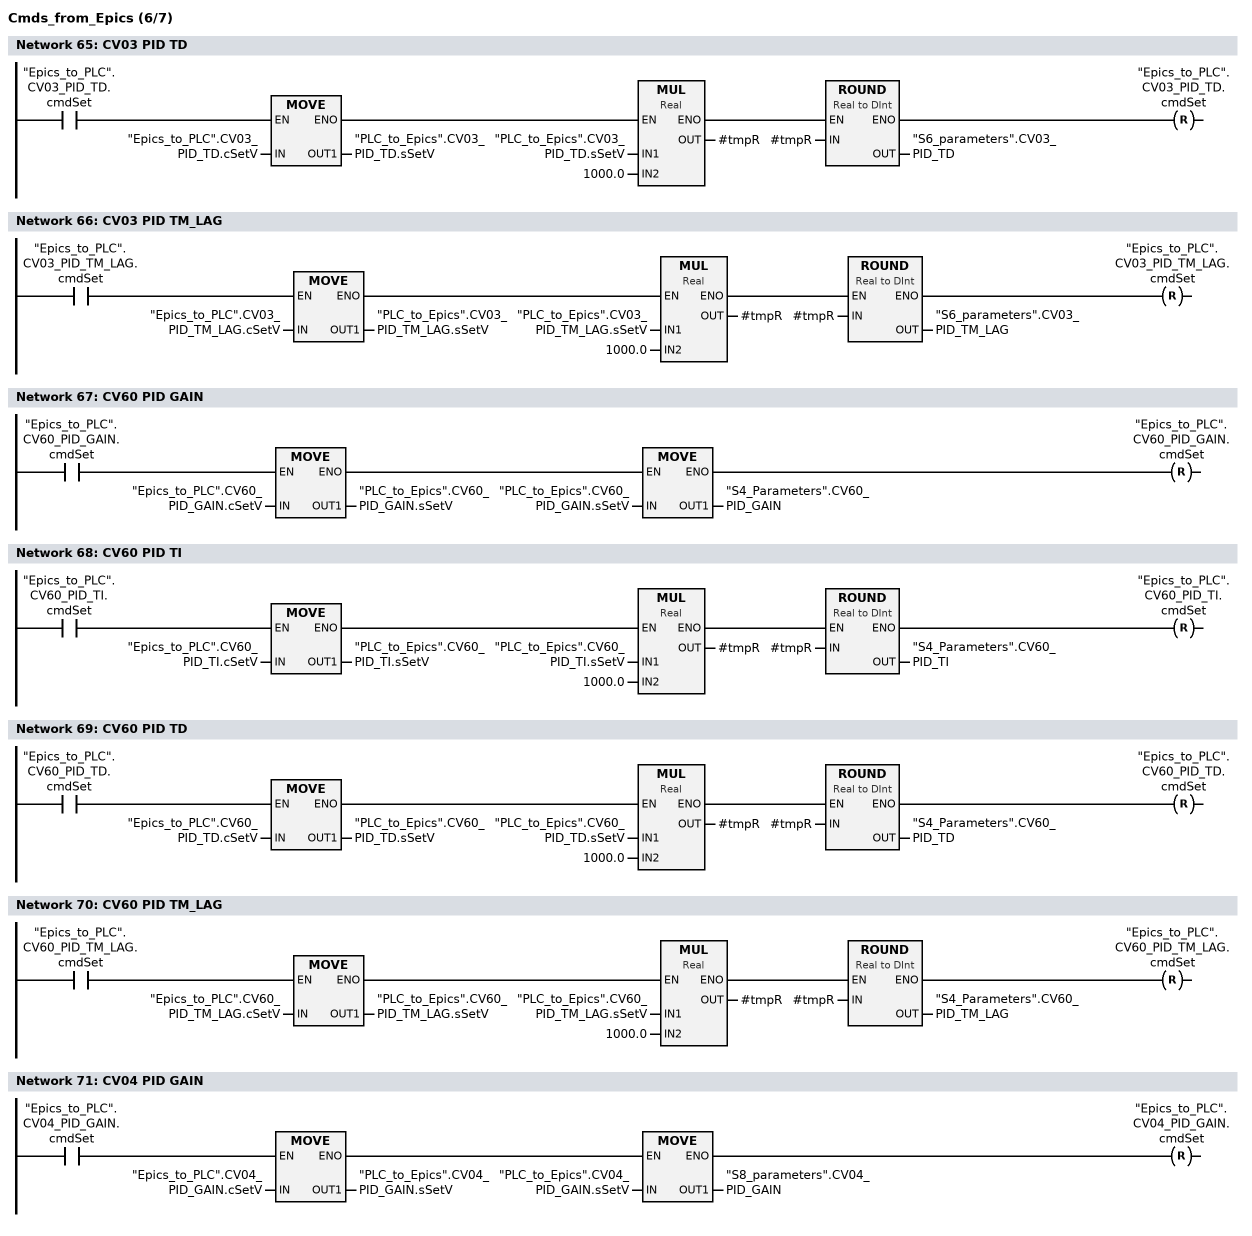
   RUNG wire#powerrail
      Contact( "Epics_to_PLC".CV03_PID_TD.cmdSet )
      { S7_GenerateENO := "TRUE" } Move(in := "Epics_to_PLC".CV03_PID_TD.cSetV, out1 => "PLC_to_Epics".CV03_PID_TD.sSetV)
      { S7_Templates := "SrcType := Real"; S7_GenerateENO := "TRUE" } Mul(in1 := "PLC_to_Epics".CV03_PID_TD.sSetV, in2 := 1000.0, out => #tmpR)
      { S7_Templates := "[SrcType := Real, DestType := DInt]"; S7_GenerateENO := "TRUE" } Round(in := #tmpR, out => "S6_parameters".CV03_PID_TD)
      R_Coil( "Epics_to_PLC".CV03_PID_TD.cmdSet )
   END_RUNG
   // the same network as SCL:
   // ENO of a box is taken as its EN; it also drops when the box reports an error
   IF "Epics_to_PLC".CV03_PID_TD.cmdSet THEN
       "PLC_to_Epics".CV03_PID_TD.sSetV := "Epics_to_PLC".CV03_PID_TD.cSetV;
       #tmpR := "PLC_to_Epics".CV03_PID_TD.sSetV * 1000.0;
       "S6_parameters".CV03_PID_TD := ROUND(#tmpR);
       "Epics_to_PLC".CV03_PID_TD.cmdSet := FALSE;
   END_IF;
END_REGION

REGION Network 66: CV03 PID TM_LAG
   RUNG wire#powerrail
      Contact( "Epics_to_PLC".CV03_PID_TM_LAG.cmdSet )
      { S7_GenerateENO := "TRUE" } Move(in := "Epics_to_PLC".CV03_PID_TM_LAG.cSetV, out1 => "PLC_to_Epics".CV03_PID_TM_LAG.sSetV)
      { S7_Templates := "SrcType := Real"; S7_GenerateENO := "TRUE" } Mul(in1 := "PLC_to_Epics".CV03_PID_TM_LAG.sSetV, in2 := 1000.0, out => #tmpR)
      { S7_Templates := "[SrcType := Real, DestType := DInt]"; S7_GenerateENO := "TRUE" } Round(in := #tmpR, out => "S6_parameters".CV03_PID_TM_LAG)
      R_Coil( "Epics_to_PLC".CV03_PID_TM_LAG.cmdSet )
   END_RUNG
   // the same network as SCL:
   // ENO of a box is taken as its EN; it also drops when the box reports an error
   IF "Epics_to_PLC".CV03_PID_TM_LAG.cmdSet THEN
       "PLC_to_Epics".CV03_PID_TM_LAG.sSetV := "Epics_to_PLC".CV03_PID_TM_LAG.cSetV;
       #tmpR := "PLC_to_Epics".CV03_PID_TM_LAG.sSetV * 1000.0;
       "S6_parameters".CV03_PID_TM_LAG := ROUND(#tmpR);
       "Epics_to_PLC".CV03_PID_TM_LAG.cmdSet := FALSE;
   END_IF;
END_REGION

REGION Network 67: CV60 PID GAIN
   RUNG wire#powerrail
      Contact( "Epics_to_PLC".CV60_PID_GAIN.cmdSet )
      { S7_GenerateENO := "TRUE" } Move(in := "Epics_to_PLC".CV60_PID_GAIN.cSetV, out1 => "PLC_to_Epics".CV60_PID_GAIN.sSetV)
      { S7_GenerateENO := "TRUE" } Move(in := "PLC_to_Epics".CV60_PID_GAIN.sSetV, out1 => "S4_Parameters".CV60_PID_GAIN)
      R_Coil( "Epics_to_PLC".CV60_PID_GAIN.cmdSet )
   END_RUNG
   // the same network as SCL:
   // ENO of a box is taken as its EN; it also drops when the box reports an error
   IF "Epics_to_PLC".CV60_PID_GAIN.cmdSet THEN
       "PLC_to_Epics".CV60_PID_GAIN.sSetV := "Epics_to_PLC".CV60_PID_GAIN.cSetV;
       "S4_Parameters".CV60_PID_GAIN := "PLC_to_Epics".CV60_PID_GAIN.sSetV;
       "Epics_to_PLC".CV60_PID_GAIN.cmdSet := FALSE;
   END_IF;
END_REGION

REGION Network 68: CV60 PID TI
   RUNG wire#powerrail
      Contact( "Epics_to_PLC".CV60_PID_TI.cmdSet )
      { S7_GenerateENO := "TRUE" } Move(in := "Epics_to_PLC".CV60_PID_TI.cSetV, out1 => "PLC_to_Epics".CV60_PID_TI.sSetV)
      { S7_Templates := "SrcType := Real"; S7_GenerateENO := "TRUE" } Mul(in1 := "PLC_to_Epics".CV60_PID_TI.sSetV, in2 := 1000.0, out => #tmpR)
      { S7_Templates := "[SrcType := Real, DestType := DInt]"; S7_GenerateENO := "TRUE" } Round(in := #tmpR, out => "S4_Parameters".CV60_PID_TI)
      R_Coil( "Epics_to_PLC".CV60_PID_TI.cmdSet )
   END_RUNG
   // the same network as SCL:
   // ENO of a box is taken as its EN; it also drops when the box reports an error
   IF "Epics_to_PLC".CV60_PID_TI.cmdSet THEN
       "PLC_to_Epics".CV60_PID_TI.sSetV := "Epics_to_PLC".CV60_PID_TI.cSetV;
       #tmpR := "PLC_to_Epics".CV60_PID_TI.sSetV * 1000.0;
       "S4_Parameters".CV60_PID_TI := ROUND(#tmpR);
       "Epics_to_PLC".CV60_PID_TI.cmdSet := FALSE;
   END_IF;
END_REGION

REGION Network 69: CV60 PID TD
   RUNG wire#powerrail
      Contact( "Epics_to_PLC".CV60_PID_TD.cmdSet )
      { S7_GenerateENO := "TRUE" } Move(in := "Epics_to_PLC".CV60_PID_TD.cSetV, out1 => "PLC_to_Epics".CV60_PID_TD.sSetV)
      { S7_Templates := "SrcType := Real"; S7_GenerateENO := "TRUE" } Mul(in1 := "PLC_to_Epics".CV60_PID_TD.sSetV, in2 := 1000.0, out => #tmpR)
      { S7_Templates := "[SrcType := Real, DestType := DInt]"; S7_GenerateENO := "TRUE" } Round(in := #tmpR, out => "S4_Parameters".CV60_PID_TD)
      R_Coil( "Epics_to_PLC".CV60_PID_TD.cmdSet )
   END_RUNG
   // the same network as SCL:
   // ENO of a box is taken as its EN; it also drops when the box reports an error
   IF "Epics_to_PLC".CV60_PID_TD.cmdSet THEN
       "PLC_to_Epics".CV60_PID_TD.sSetV := "Epics_to_PLC".CV60_PID_TD.cSetV;
       #tmpR := "PLC_to_Epics".CV60_PID_TD.sSetV * 1000.0;
       "S4_Parameters".CV60_PID_TD := ROUND(#tmpR);
       "Epics_to_PLC".CV60_PID_TD.cmdSet := FALSE;
   END_IF;
END_REGION

REGION Network 70: CV60 PID TM_LAG
   RUNG wire#powerrail
      Contact( "Epics_to_PLC".CV60_PID_TM_LAG.cmdSet )
      { S7_GenerateENO := "TRUE" } Move(in := "Epics_to_PLC".CV60_PID_TM_LAG.cSetV, out1 => "PLC_to_Epics".CV60_PID_TM_LAG.sSetV)
      { S7_Templates := "SrcType := Real"; S7_GenerateENO := "TRUE" } Mul(in1 := "PLC_to_Epics".CV60_PID_TM_LAG.sSetV, in2 := 1000.0, out => #tmpR)
      { S7_Templates := "[SrcType := Real, DestType := DInt]"; S7_GenerateENO := "TRUE" } Round(in := #tmpR, out => "S4_Parameters".CV60_PID_TM_LAG)
      R_Coil( "Epics_to_PLC".CV60_PID_TM_LAG.cmdSet )
   END_RUNG
   // the same network as SCL:
   // ENO of a box is taken as its EN; it also drops when the box reports an error
   IF "Epics_to_PLC".CV60_PID_TM_LAG.cmdSet THEN
       "PLC_to_Epics".CV60_PID_TM_LAG.sSetV := "Epics_to_PLC".CV60_PID_TM_LAG.cSetV;
       #tmpR := "PLC_to_Epics".CV60_PID_TM_LAG.sSetV * 1000.0;
       "S4_Parameters".CV60_PID_TM_LAG := ROUND(#tmpR);
       "Epics_to_PLC".CV60_PID_TM_LAG.cmdSet := FALSE;
   END_IF;
END_REGION

REGION Network 71: CV04 PID GAIN
   RUNG wire#powerrail
      Contact( "Epics_to_PLC".CV04_PID_GAIN.cmdSet )
      { S7_GenerateENO := "TRUE" } Move(in := "Epics_to_PLC".CV04_PID_GAIN.cSetV, out1 => "PLC_to_Epics".CV04_PID_GAIN.sSetV)
      { S7_GenerateENO := "TRUE" } Move(in := "PLC_to_Epics".CV04_PID_GAIN.sSetV, out1 => "S8_parameters".CV04_PID_GAIN)
      R_Coil( "Epics_to_PLC".CV04_PID_GAIN.cmdSet )
   END_RUNG
   // the same network as SCL:
   // ENO of a box is taken as its EN; it also drops when the box reports an error
   IF "Epics_to_PLC".CV04_PID_GAIN.cmdSet THEN
       "PLC_to_Epics".CV04_PID_GAIN.sSetV := "Epics_to_PLC".CV04_PID_GAIN.cSetV;
       "S8_parameters".CV04_PID_GAIN := "PLC_to_Epics".CV04_PID_GAIN.sSetV;
       "Epics_to_PLC".CV04_PID_GAIN.cmdSet := FALSE;
   END_IF;
END_REGION

REGION Network 72: CV04 PID TI